   "DB_HMI_ARG1_Seq1_DelaySelect_Blue{4}" : Bool = PLC DB_HMI.ARG1_Seq1_DelaySelect_Blue[4] AT %DB1.DBX0.0, 100 ms
   "DB_HMI_ARG1_Seq1_DelaySelect_Blue{5}" : Bool = PLC DB_HMI.ARG1_Seq1_DelaySelect_Blue[5] AT %DB1.DBX0.0, 100 ms
   "DB_HMI_ARG1_Seq1_DelaySelect_Blue{6}" : Bool = PLC DB_HMI.ARG1_Seq1_DelaySelect_Blue[6] AT %DB1.DBX0.0, 100 ms
   "DB_HMI_ARG1_Seq1_DelaySelect_Blue{7}" : Bool = PLC DB_HMI.ARG1_Seq1_DelaySelect_Blue[7] AT %DB1.DBX0.0, 100 ms
   "DB_HMI_ARG1_Seq1_DelaySelect_Blue{8}" : Bool = PLC DB_HMI.ARG1_Seq1_DelaySelect_Blue[8] AT %DB1.DBX0.0, 100 ms
   "DB_HMI_ARG1_Seq1_DelaySelect_Blue{9}" : Bool = PLC DB_HMI.ARG1_Seq1_DelaySelect_Blue[9] AT %DB1.DBX0.0, 100 ms
   "DB_HMI_ARG1_Seq1_DelaySelect_Blue{10}" : Bool = PLC DB_HMI.ARG1_Seq1_DelaySelect_Blue[10] AT %DB1.DBX0.0, 100 ms
   "DB_HMI_Global_Cmd_Auto" : Bool = PLC DB_HMI.Global_Cmd_Auto, 100 ms
   "DB_HMI_Global_Cmd_Man" : Bool = PLC DB_HMI.Global_Cmd_Man, 100 ms
   "DB_HMI_Global_Cmd_Start" : Bool = PLC DB_HMI.Global_Cmd_Start, 100 ms
   "DB_HMI_Global_Cmd_Stop" : Bool = PLC DB_HMI.Global_Cmd_Stop, 100 ms
   "DB_HMI_Global_Status_Man" : Bool = PLC DB_HMI.Global_Status_Man AT %DB1.DBW0, 100 ms
   "DB_HMI_Global_Status_Auto" : Bool = PLC DB_HMI.Global_Status_Auto AT %DB1.DBW0, 100 ms
   "DB_HMI_Global_selection" : Int = PLC DB_HMI.Global_selection AT %DB1.DBW0, 100 ms
   "DB_HMI_inProduction" : Int = PLC DB_HMI.ARG1_Seq1_inProduction AT %DB1.DBW0, 100 ms

HMI tags "PLC_2_tags"
   "DB_HMI_ARG1_Seq1_S1(1)" : Bool = PLC DB_HMI.ARG1_Seq1_S1, 100 ms
   "DB_HMI_ARG1_Seq1_T1(1)" : Bool = PLC DB_HMI.ARG1_Seq1_T1, 100 ms
   "DB_HMI_ARG1_Seq1_S2(1)" : Bool = PLC DB_HMI.ARG1_Seq1_S2, 100 ms
   "DB_HMI_ARG1_Seq1_T2(1)" : Bool = PLC DB_HMI.ARG1_Seq1_T2, 100 ms
   "DB_HMI_ARG1_Seq1_S3(1)" : Bool = PLC DB_HMI.ARG1_Seq1_S3, 100 ms
   "DB_HMI_ARG1_Seq1_T3(1)" : Bool = PLC DB_HMI.ARG1_Seq1_T3, 100 ms
   "DB_HMI_ARG1_Seq1_S4(1)" : Bool = PLC DB_HMI.ARG1_Seq1_S4, 100 ms
   "DB_HMI_ARG1_Seq1_T4(1)" : Bool = PLC DB_HMI.ARG1_Seq1_T4, 100 ms
   "DB_HMI_ARG1_Seq1_S5(1)" : Bool = PLC DB_HMI.ARG1_Seq1_S5, 100 ms
   "DB_HMI_ARG1_Seq1_T5(1)" : Bool = PLC DB_HMI.ARG1_Seq1_T5, 100 ms
   "DB_HMI_ARG1_Seq1_S6(1)" : Bool = PLC DB_HMI.ARG1_Seq1_S6, 100 ms
   "DB_HMI_ARG1_Seq1_T6(1)" : Bool = PLC DB_HMI.ARG1_Seq1_T6, 100 ms
   "DB_HMI_ARG1_Seq1_S7(1)" : Bool = PLC DB_HMI.ARG1_Seq1_S7, 100 ms
   "DB_HMI_ARG1_Seq1_T7(1)" : Bool = PLC DB_HMI.ARG1_Seq1_T7, 100 ms
   "DB_HMI_ARG1_Seq1_S8(1)" : Bool = PLC DB_HMI.ARG1_Seq1_S8, 100 ms
   "DB_HMI_ARG1_Seq1_T8(1)" : Bool = PLC DB_HMI.ARG1_Seq1_T8, 100 ms
   "DB_HMI_ARG1_Seq1_S9(1)" : Bool = PLC DB_HMI.ARG1_Seq1_S9, 100 ms
   "DB_HMI_ARG1_Seq1_T9(1)" : Bool = PLC DB_HMI.ARG1_Seq1_T9, 100 ms
   "DB_HMI_ARG1_Seq1_S10(1)" : Bool = PLC DB_HMI.ARG1_Seq1_S10, 100 ms
   "DB_HMI_ARG1_Seq1_T10(1)" : Bool = PLC DB_HMI.ARG1_Seq1_T10, 100 ms
   "DB_HMI_ARG1_Seq1_S11(1)" : Bool = PLC DB_HMI.ARG1_Seq1_S11, 100 ms
   "DB_HMI_ARG1_Seq1_T11(1)" : Bool = PLC DB_HMI.ARG1_Seq1_T11, 100 ms
   "DB_HMI_ARG1_Seq1_S12(1)" : Bool = PLC DB_HMI.ARG1_Seq1_S12, 100 ms
   "DB_HMI_ARG1_Seq1_T12(1)" : Bool = PLC DB_HMI.ARG1_Seq1_T12, 100 ms
   "DB_HMI_ARG1_Seq1_S13(1)" : Bool = PLC DB_HMI.ARG1_Seq1_S13, 100 ms
   "DB_HMI_ARG1_Seq1_T13(1)" : Bool = PLC DB_HMI.ARG1_Seq1_T13, 100 ms
   "DB_HMI_ARG1_Seq1_S14(1)" : Bool = PLC DB_HMI.ARG1_Seq1_S14, 100 ms
   "DB_HMI_ARG1_Seq1_T14(1)" : Bool = PLC DB_HMI.ARG1_Seq1_T14, 100 ms
   "DB_HMI_ARG1_Seq1_S15(1)" : Bool = PLC DB_HMI.ARG1_Seq1_S15, 100 ms
   "DB_HMI_ARG1_Seq1_T15(1)" : Bool = PLC DB_HMI.ARG1_Seq1_T15, 100 ms
   "DB_HMI_ARG1_Seq1_S16(1)" : Bool = PLC DB_HMI.ARG1_Seq1_S16, 100 ms
   "DB_HMI_ARG1_Seq1_T16(1)" : Bool = PLC DB_HMI.ARG1_Seq1_T16, 100 ms
   "DB_HMI_ARG1_Seq1_S17(1)" : Bool = PLC DB_HMI.ARG1_Seq1_S17, 100 ms
   "DB_HMI_ARG1_Seq1_T17(1)" : Bool = PLC DB_HMI.ARG1_Seq1_T17, 100 ms
   "DB_HMI_ARG1_Seq1_S18(1)" : Bool = PLC DB_HMI.ARG1_Seq1_S18, 100 ms
   "DB_HMI_ARG1_Seq1_T18(1)" : Bool = PLC DB_HMI.ARG1_Seq1_T18, 100 ms
   "DB_HMI_ARG1_Seq1_S19(1)" : Bool = PLC DB_HMI.ARG1_Seq1_S19, 100 ms
   "DB_HMI_ARG1_Seq1_T19(1)" : Bool = PLC DB_HMI.ARG1_Seq1_T19, 100 ms
   "DB_HMI_inputTimes(1)" : Array [0..8] of DInt = PLC DB_HMI.inputTimes, 100 ms
   "DB_HMI_dropdown_selection(1)" : Int = PLC DB_HMI.dropdown_selection, 100 ms
   "DB_HMI_ARG1_Seq1_Status_Idle(1)" : Bool = PLC DB_HMI.ARG1_Seq1_Status_Idle, 100 ms
   "DB_HMI_ARG1_Seq1_Status_Busy(1)" : Bool = PLC DB_HMI.ARG1_Seq1_Status_Busy, 100 ms
   "DB_HMI_ARG1_Seq1_Status_Man(1)" : Bool = PLC DB_HMI.ARG1_Seq1_Status_Man, 100 ms
   "DB_HMI_ARG1_Seq1_Status_Auto(1)" : Bool = PLC DB_HMI.ARG1_Seq1_Status_Auto, 100 ms
   "DB_HMI_ARG1_Seq1_Cmd_Man(1)" : Bool = PLC DB_HMI.ARG1_Seq1_Cmd_Man, 100 ms
   "DB_HMI_ARG1_Seq1_Cmd_Auto(1)" : Bool = PLC DB_HMI.ARG1_Seq1_Cmd_Auto, 100 ms
   "DB_HMI_ARG1_Seq1_Cmd_Stop(1)" : Bool = PLC DB_HMI.ARG1_Seq1_Cmd_Stop, 100 ms
   "DB_HMI_ARG1_Seq1_Cmd_Start(1)" : Bool = PLC DB_HMI.ARG1_Seq1_Cmd_Start, 100 ms
   "DB_HMI_ARG1_Seq1_Cmd_DelayReset(1)" : Bool = PLC DB_HMI.ARG1_Seq1_Cmd_DelayReset, 100 ms
   "DB_HMI_ARG1_Seq1_Calculated_PT_Red(1)" : Time = PLC DB_HMI.ARG1_Seq1_Calculated_PT_Red, 100 ms
   "DB_HMI_ARG1_Seq1_Calculated_PT_Green(1)" : Time = PLC DB_HMI.ARG1_Seq1_Calculated_PT_Green, 100 ms
   "DB_HMI_ARG1_Seq1_Calculated_PT_Blue(1)" : Time = PLC DB_HMI.ARG1_Seq1_Calculated_PT_Blue, 100 ms
   "DB_HMI_ARG1_Seq1_Messured_PT_Red(1)" : Time = PLC DB_HMI.ARG1_Seq1_Messured_PT_Red, 100 ms
   "DB_HMI_ARG1_Seq1_Messured_PT_Green(1)" : Time = PLC DB_HMI.ARG1_Seq1_Messured_PT_Green, 100 ms
   "DB_HMI_ARG1_Seq1_Messured_PT_Blue(1)" : Time = PLC DB_HMI.ARG1_Seq1_Messured_PT_Blue, 100 ms
   "DB_HMI_ARG1_Seq1_DelaySelect_Red(1)" : Array [0..8] of Bool = PLC DB_HMI.ARG1_Seq1_DelaySelect_Red, 100 ms
   "DB_HMI_ARG1_Seq1_DelaySelect_Green(1)" : Array [0..8] of Bool = PLC DB_HMI.ARG1_Seq1_DelaySelect_Green, 100 ms
   "DB_HMI_ARG1_Seq1_DelaySelect_Blue(1)" : Array [0..8] of Bool = PLC DB_HMI.ARG1_Seq1_DelaySelect_Blue, 100 ms
   "DB_HMI_ARG1_Seq1_DelaySelect_Red{2}(1)" : Bool = PLC DB_HMI.ARG1_Seq1_DelaySelect_Red[2] AT %DB1.DBW0, 100 ms
   "DB_HMI_ARG1_Seq1_DelaySelect_Red{3}(1)" : Bool = PLC DB_HMI.ARG1_Seq1_DelaySelect_Red[3] AT %DB1.DBW0, 100 ms
   "DB_HMI_ARG1_Seq1_DelaySelect_Red{4}(1)" : Bool = PLC DB_HMI.ARG1_Seq1_DelaySelect_Red[4] AT %DB1.DBW0, 100 ms
   "DB_HMI_ARG1_Seq1_DelaySelect_Red{5}(1)" : Bool = PLC DB_HMI.ARG1_Seq1_DelaySelect_Red[5] AT %DB1.DBW0, 100 ms
   "DB_HMI_ARG1_Seq1_DelaySelect_Red{6}(1)" : Bool = PLC DB_HMI.ARG1_Seq1_DelaySelect_Red[6] AT %DB1.DBW0, 100 ms
   "DB_HMI_ARG1_Seq1_DelaySelect_Red{7}(1)" : Bool = PLC DB_HMI.ARG1_Seq1_DelaySelect_Red[7] AT %DB1.DBW0, 100 ms
   "DB_HMI_ARG1_Seq1_DelaySelect_Red{8}(1)" : Bool = PLC DB_HMI.ARG1_Seq1_DelaySelect_Red[8] AT %DB1.DBW0, 100 ms
   "DB_HMI_ARG1_Seq1_DelaySelect_Red{9}(1)" : Bool = PLC DB_HMI.ARG1_Seq1_DelaySelect_Red[9] AT %DB1.DBW0, 100 ms
   "DB_HMI_ARG1_Seq1_DelaySelect_Red{10}(1)" : Bool = PLC DB_HMI.ARG1_Seq1_DelaySelect_Red[10] AT %DB1.DBW0, 100 ms
   "DB_HMI_ARG1_Seq1_DelaySelect_Green{2}(1)" : Bool = PLC DB_HMI.ARG1_Seq1_DelaySelect_Green[2] AT %DB1.DBX0.0, 100 ms
   "DB_HMI_ARG1_Seq1_DelaySelect_Green{3}(1)" : Bool = PLC DB_HMI.ARG1_Seq1_DelaySelect_Green[3] AT %DB1.DBX0.0, 100 ms
   "DB_HMI_ARG1_Seq1_DelaySelect_Green{4}(1)" : Bool = PLC DB_HMI.ARG1_Seq1_DelaySelect_Green[4] AT %DB1.DBX0.0, 100 ms
   "DB_HMI_ARG1_Seq1_DelaySelect_Green{5}(1)" : Bool = PLC DB_HMI.ARG1_Seq1_DelaySelect_Green[5] AT %DB1.DBX0.0, 100 ms
   "DB_HMI_ARG1_Seq1_DelaySelect_Green{6}(1)" : Bool = PLC DB_HMI.ARG1_Seq1_DelaySelect_Green[6] AT %DB1.DBX0.0, 100 ms
   "DB_HMI_ARG1_Seq1_DelaySelect_Green{7}(1)" : Bool = PLC DB_HMI.ARG1_Seq1_DelaySelect_Green[7] AT %DB1.DBX0.0, 100 ms
   "DB_HMI_ARG1_Seq1_DelaySelect_Green{8}(1)" : Bool = PLC DB_HMI.ARG1_Seq1_DelaySelect_Green[8] AT %DB1.DBX0.0, 100 ms
   "DB_HMI_ARG1_Seq1_DelaySelect_Green{9}(1)" : Bool = PLC DB_HMI.ARG1_Seq1_DelaySelect_Green[9] AT %DB1.DBX0.0, 100 ms
   "DB_HMI_ARG1_Seq1_DelaySelect_Green{10}(1)" : Bool = PLC DB_HMI.ARG1_Seq1_DelaySelect_Green[10] AT %DB1.DBX0.0, 100 ms
   "DB_HMI_ARG1_Seq1_DelaySelect_Blue{2}(1)" : Bool = PLC DB_HMI.ARG1_Seq1_DelaySelect_Blue[2] AT %DB1.DBX0.0, 100 ms
   "DB_HMI_ARG1_Seq1_DelaySelect_Blue{3}(1)" : Bool = PLC DB_HMI.ARG1_Seq1_DelaySelect_Blue[3] AT %DB1.DBX0.0, 100 ms
   "DB_HMI_ARG1_Seq1_DelaySelect_Blue{4}(1)" : Bool = PLC DB_HMI.ARG1_Seq1_DelaySelect_Blue[4] AT %DB1.DBX0.0, 100 ms
   "DB_HMI_ARG1_Seq1_DelaySelect_Blue{5}(1)" : Bool = PLC DB_HMI.ARG1_Seq1_DelaySelect_Blue[5] AT %DB1.DBX0.0, 100 ms
   "DB_HMI_ARG1_Seq1_DelaySelect_Blue{6}(1)" : Bool = PLC DB_HMI.ARG1_Seq1_DelaySelect_Blue[6] AT %DB1.DBX0.0, 100 ms
   "DB_HMI_ARG1_Seq1_DelaySelect_Blue{7}(1)" : Bool = PLC DB_HMI.ARG1_Seq1_DelaySelect_Blue[7] AT %DB1.DBX0.0, 100 ms
   "DB_HMI_ARG1_Seq1_DelaySelect_Blue{8}(1)" : Bool = PLC DB_HMI.ARG1_Seq1_DelaySelect_Blue[8] AT %DB1.DBX0.0, 100 ms
   "DB_HMI_ARG1_Seq1_DelaySelect_Blue{9}(1)" : Bool = PLC DB_HMI.ARG1_Seq1_DelaySelect_Blue[9] AT %DB1.DBX0.0, 100 ms
   "DB_HMI_ARG1_Seq1_DelaySelect_Blue{10}(1)" : Bool = PLC DB_HMI.ARG1_Seq1_DelaySelect_Blue[10] AT %DB1.DBX0.0, 100 ms
   "DB_HMI_Global_Cmd_Auto(1)" : Bool = PLC DB_HMI.Global_Cmd_Auto, 100 ms
   "DB_HMI_Global_Cmd_Man(1)" : Bool = PLC DB_HMI.Global_Cmd_Man, 100 ms
   "DB_HMI_Global_Cmd_Start(1)" : Bool = PLC DB_HMI.Global_Cmd_Start, 100 ms
   "DB_HMI_Global_Cmd_Stop(1)" : Bool = PLC DB_HMI.Global_Cmd_Stop, 100 ms
   "DB_HMI_inProduction(1)" : Int = PLC DB_HMI.ARG1_Seq1_inProduction AT %DB1.DBW0, 100 ms

HMI tags "PLC_3_tags"
   "DB_HMI_ARG1_Seq1_S1(2)" : Bool = PLC DB_HMI.ARG1_Seq1_S1, 100 ms
   "DB_HMI_ARG1_Seq1_T1(2)" : Bool = PLC DB_HMI.ARG1_Seq1_T1, 100 ms
   "DB_HMI_ARG1_Seq1_S2(2)" : Bool = PLC DB_HMI.ARG1_Seq1_S2, 100 ms
   "DB_HMI_ARG1_Seq1_T2(2)" : Bool = PLC DB_HMI.ARG1_Seq1_T2, 100 ms
   "DB_HMI_ARG1_Seq1_S3(2)" : Bool = PLC DB_HMI.ARG1_Seq1_S3, 100 ms
   "DB_HMI_ARG1_Seq1_T3(2)" : Bool = PLC DB_HMI.ARG1_Seq1_T3, 100 ms
   "DB_HMI_ARG1_Seq1_S4(2)" : Bool = PLC DB_HMI.ARG1_Seq1_S4, 100 ms
   "DB_HMI_ARG1_Seq1_T4(2)" : Bool = PLC DB_HMI.ARG1_Seq1_T4, 100 ms
   "DB_HMI_ARG1_Seq1_S5(2)" : Bool = PLC DB_HMI.ARG1_Seq1_S5, 100 ms
   "DB_HMI_ARG1_Seq1_T5(2)" : Bool = PLC DB_HMI.ARG1_Seq1_T5, 100 ms
   "DB_HMI_ARG1_Seq1_S6(2)" : Bool = PLC DB_HMI.ARG1_Seq1_S6, 100 ms
   "DB_HMI_ARG1_Seq1_T6(2)" : Bool = PLC DB_HMI.ARG1_Seq1_T6, 100 ms
   "DB_HMI_ARG1_Seq1_S7(2)" : Bool = PLC DB_HMI.ARG1_Seq1_S7, 100 ms
   "DB_HMI_ARG1_Seq1_T7(2)" : Bool = PLC DB_HMI.ARG1_Seq1_T7, 100 ms
   "DB_HMI_ARG1_Seq1_S8(2)" : Bool = PLC DB_HMI.ARG1_Seq1_S8, 100 ms
   "DB_HMI_ARG1_Seq1_T8(2)" : Bool = PLC DB_HMI.ARG1_Seq1_T8, 100 ms
   "DB_HMI_ARG1_Seq1_S9(2)" : Bool = PLC DB_HMI.ARG1_Seq1_S9, 100 ms
   "DB_HMI_ARG1_Seq1_T9(2)" : Bool = PLC DB_HMI.ARG1_Seq1_T9, 100 ms
   "DB_HMI_ARG1_Seq1_S10(2)" : Bool = PLC DB_HMI.ARG1_Seq1_S10, 100 ms
   "DB_HMI_ARG1_Seq1_T10(2)" : Bool = PLC DB_HMI.ARG1_Seq1_T10, 100 ms
   "DB_HMI_ARG1_Seq1_S11(2)" : Bool = PLC DB_HMI.ARG1_Seq1_S11, 100 ms
   "DB_HMI_ARG1_Seq1_T11(2)" : Bool = PLC DB_HMI.ARG1_Seq1_T11, 100 ms
   "DB_HMI_ARG1_Seq1_S12(2)" : Bool = PLC DB_HMI.ARG1_Seq1_S12, 100 ms
   "DB_HMI_ARG1_Seq1_T12(2)" : Bool = PLC DB_HMI.ARG1_Seq1_T12, 100 ms
   "DB_HMI_ARG1_Seq1_S13(2)" : Bool = PLC DB_HMI.ARG1_Seq1_S13, 100 ms
   "DB_HMI_ARG1_Seq1_T13(2)" : Bool = PLC DB_HMI.ARG1_Seq1_T13, 100 ms
   "DB_HMI_ARG1_Seq1_S14(2)" : Bool = PLC DB_HMI.ARG1_Seq1_S14, 100 ms
   "DB_HMI_ARG1_Seq1_T14(2)" : Bool = PLC DB_HMI.ARG1_Seq1_T14, 100 ms
   "DB_HMI_ARG1_Seq1_S15(2)" : Bool = PLC DB_HMI.ARG1_Seq1_S15, 100 ms
   "DB_HMI_ARG1_Seq1_T15(2)" : Bool = PLC DB_HMI.ARG1_Seq1_T15, 100 ms
   "DB_HMI_ARG1_Seq1_S16(2)" : Bool = PLC DB_HMI.ARG1_Seq1_S16, 100 ms
   "DB_HMI_ARG1_Seq1_T16(2)" : Bool = PLC DB_HMI.ARG1_Seq1_T16, 100 ms
   "DB_HMI_ARG1_Seq1_S17(2)" : Bool = PLC DB_HMI.ARG1_Seq1_S17, 100 ms
   "DB_HMI_ARG1_Seq1_T17(2)" : Bool = PLC DB_HMI.ARG1_Seq1_T17, 100 ms
   "DB_HMI_ARG1_Seq1_S18(2)" : Bool = PLC DB_HMI.ARG1_Seq1_S18, 100 ms
   "DB_HMI_ARG1_Seq1_T18(2)" : Bool = PLC DB_HMI.ARG1_Seq1_T18, 100 ms
   "DB_HMI_ARG1_Seq1_S19(2)" : Bool = PLC DB_HMI.ARG1_Seq1_S19, 100 ms
   "DB_HMI_ARG1_Seq1_T19(2)" : Bool = PLC DB_HMI.ARG1_Seq1_T19, 100 ms
   "DB_HMI_inputTimes(2)" : Array [0..8] of DInt = PLC DB_HMI.inputTimes, 100 ms
   "DB_HMI_dropdown_selection(2)" : Int = PLC DB_HMI.dropdown_selection, 100 ms
   "DB_HMI_ARG1_Seq1_Status_Idle(2)" : Bool = PLC DB_HMI.ARG1_Seq1_Status_Idle, 100 ms
   "DB_HMI_ARG1_Seq1_Status_Busy(2)" : Bool = PLC DB_HMI.ARG1_Seq1_Status_Busy, 100 ms
   "DB_HMI_ARG1_Seq1_Status_Man(2)" : Bool = PLC DB_HMI.ARG1_Seq1_Status_Man, 100 ms
   "DB_HMI_ARG1_Seq1_Status_Auto(2)" : Bool = PLC DB_HMI.ARG1_Seq1_Status_Auto, 100 ms
   "DB_HMI_ARG1_Seq1_Cmd_Man(2)" : Bool = PLC DB_HMI.ARG1_Seq1_Cmd_Man, 100 ms
   "DB_HMI_ARG1_Seq1_Cmd_Auto(2)" : Bool = PLC DB_HMI.ARG1_Seq1_Cmd_Auto, 100 ms
   "DB_HMI_ARG1_Seq1_Cmd_Stop(2)" : Bool = PLC DB_HMI.ARG1_Seq1_Cmd_Stop, 100 ms
   "DB_HMI_ARG1_Seq1_Cmd_Start(2)" : Bool = PLC DB_HMI.ARG1_Seq1_Cmd_Start, 100 ms
   "DB_HMI_ARG1_Seq1_Cmd_DelayReset(2)" : Bool = PLC DB_HMI.ARG1_Seq1_Cmd_DelayReset, 100 ms
   "DB_HMI_ARG1_Seq1_Calculated_PT_Red(2)" : Time = PLC DB_HMI.ARG1_Seq1_Calculated_PT_Red, 100 ms
   "DB_HMI_ARG1_Seq1_Calculated_PT_Green(2)" : Time = PLC DB_HMI.ARG1_Seq1_Calculated_PT_Green, 100 ms
   "DB_HMI_ARG1_Seq1_Calculated_PT_Blue(2)" : Time = PLC DB_HMI.ARG1_Seq1_Calculated_PT_Blue, 100 ms
   "DB_HMI_ARG1_Seq1_Messured_PT_Red(2)" : Time = PLC DB_HMI.ARG1_Seq1_Messured_PT_Red, 100 ms
   "DB_HMI_ARG1_Seq1_Messured_PT_Green(2)" : Time = PLC DB_HMI.ARG1_Seq1_Messured_PT_Green, 100 ms
   "DB_HMI_ARG1_Seq1_Messured_PT_Blue(2)" : Time = PLC DB_HMI.ARG1_Seq1_Messured_PT_Blue, 100 ms
   "DB_HMI_ARG1_Seq1_DelaySelect_Red(2)" : Array [0..8] of Bool = PLC DB_HMI.ARG1_Seq1_DelaySelect_Red, 100 ms
   "DB_HMI_ARG1_Seq1_DelaySelect_Green(2)" : Array [0..8] of Bool = PLC DB_HMI.ARG1_Seq1_DelaySelect_Green, 100 ms
   "DB_HMI_ARG1_Seq1_DelaySelect_Blue(2)" : Array [0..8] of Bool = PLC DB_HMI.ARG1_Seq1_DelaySelect_Blue, 100 ms
   "DB_HMI_ARG1_Seq1_DelaySelect_Red{2}(2)" : Bool = PLC DB_HMI.ARG1_Seq1_DelaySelect_Red[2], 100 ms
   "DB_HMI_ARG1_Seq1_DelaySelect_Red{3}(2)" : Bool = PLC DB_HMI.ARG1_Seq1_DelaySelect_Red[3], 100 ms
   "DB_HMI_ARG1_Seq1_DelaySelect_Red{4}(2)" : Bool = PLC DB_HMI.ARG1_Seq1_DelaySelect_Red[4], 100 ms
   "DB_HMI_ARG1_Seq1_DelaySelect_Red{5}(2)" : Bool = PLC DB_HMI.ARG1_Seq1_DelaySelect_Red[5], 100 ms
   "DB_HMI_ARG1_Seq1_DelaySelect_Red{6}(2)" : Bool = PLC DB_HMI.ARG1_Seq1_DelaySelect_Red[6], 100 ms
   "DB_HMI_ARG1_Seq1_DelaySelect_Red{7}(2)" : Bool = PLC DB_HMI.ARG1_Seq1_DelaySelect_Red[7], 100 ms
   "DB_HMI_ARG1_Seq1_DelaySelect_Red{8}(2)" : Bool = PLC DB_HMI.ARG1_Seq1_DelaySelect_Red[8], 100 ms
   "DB_HMI_ARG1_Seq1_DelaySelect_Red{9}(2)" : Bool = PLC DB_HMI.ARG1_Seq1_DelaySelect_Red[9], 100 ms
   "DB_HMI_ARG1_Seq1_DelaySelect_Red{10}(2)" : Bool = PLC DB_HMI.ARG1_Seq1_DelaySelect_Red[10], 100 ms
   "DB_HMI_ARG1_Seq1_DelaySelect_Green{2}(2)" : Bool = PLC DB_HMI.ARG1_Seq1_DelaySelect_Green[2], 100 ms
   "DB_HMI_ARG1_Seq1_DelaySelect_Green{3}(2)" : Bool = PLC DB_HMI.ARG1_Seq1_DelaySelect_Green[3], 100 ms
   "DB_HMI_ARG1_Seq1_DelaySelect_Green{4}(2)" : Bool = PLC DB_HMI.ARG1_Seq1_DelaySelect_Green[4], 100 ms
   "DB_HMI_ARG1_Seq1_DelaySelect_Green{5}(2)" : Bool = PLC DB_HMI.ARG1_Seq1_DelaySelect_Green[5], 100 ms
   "DB_HMI_ARG1_Seq1_DelaySelect_Green{6}(2)" : Bool = PLC DB_HMI.ARG1_Seq1_DelaySelect_Green[6], 100 ms
   "DB_HMI_ARG1_Seq1_DelaySelect_Green{7}(2)" : Bool = PLC DB_HMI.ARG1_Seq1_DelaySelect_Green[7], 100 ms
   "DB_HMI_ARG1_Seq1_DelaySelect_Green{8}(2)" : Bool = PLC DB_HMI.ARG1_Seq1_DelaySelect_Green[8], 100 ms
   "DB_HMI_ARG1_Seq1_DelaySelect_Green{9}(2)" : Bool = PLC DB_HMI.ARG1_Seq1_DelaySelect_Green[9], 100 ms
   "DB_HMI_ARG1_Seq1_DelaySelect_Green{10}(2)" : Bool = PLC DB_HMI.ARG1_Seq1_DelaySelect_Green[10], 100 ms
   "DB_HMI_ARG1_Seq1_DelaySelect_Blue{2}(2)" : Bool = PLC DB_HMI.ARG1_Seq1_DelaySelect_Blue[2], 100 ms
   "DB_HMI_ARG1_Seq1_DelaySelect_Blue{3}(2)" : Bool = PLC DB_HMI.ARG1_Seq1_DelaySelect_Blue[3], 100 ms
   "DB_HMI_ARG1_Seq1_DelaySelect_Blue{4}(2)" : Bool = PLC DB_HMI.ARG1_Seq1_DelaySelect_Blue[4], 100 ms
   "DB_HMI_ARG1_Seq1_DelaySelect_Blue{5}(2)" : Bool = PLC DB_HMI.ARG1_Seq1_DelaySelect_Blue[5], 100 ms
   "DB_HMI_ARG1_Seq1_DelaySelect_Blue{6}(2)" : Bool = PLC DB_HMI.ARG1_Seq1_DelaySelect_Blue[6], 100 ms
   "DB_HMI_ARG1_Seq1_DelaySelect_Blue{7}(2)" : Bool = PLC DB_HMI.ARG1_Seq1_DelaySelect_Blue[7], 100 ms
   "DB_HMI_ARG1_Seq1_DelaySelect_Blue{8}(2)" : Bool = PLC DB_HMI.ARG1_Seq1_DelaySelect_Blue[8], 100 ms
   "DB_HMI_ARG1_Seq1_DelaySelect_Blue{9}(2)" : Bool = PLC DB_HMI.ARG1_Seq1_DelaySelect_Blue[9], 100 ms
   "DB_HMI_ARG1_Seq1_DelaySelect_Blue{10}(2)" : Bool = PLC DB_HMI.ARG1_Seq1_DelaySelect_Blue[10], 100 ms
   "DB_HMI_Global_Cmd_Auto(2)" : Bool = PLC DB_HMI.Global_Cmd_Auto, 100 ms
   "DB_HMI_Global_Cmd_Man(2)" : Bool = PLC DB_HMI.Global_Cmd_Man, 100 ms
   "DB_HMI_Global_Cmd_Start(2)" : Bool = PLC DB_HMI.Global_Cmd_Start, 100 ms
   "DB_HMI_Global_Cmd_Stop(2)" : Bool = PLC DB_HMI.Global_Cmd_Stop, 100 ms
   "DB_HMI_inProduction(2)" : Int = PLC DB_HMI.ARG1_Seq1_inProduction AT %DB1.DBW0, 100 ms

HMI tags "PLC_4_tags"
   "DB_HMI_ARG1_Seq1_S1(3)" : Bool = PLC DB_HMI.ARG1_Seq1_S1, 100 ms
   "DB_HMI_ARG1_Seq1_T1(3)" : Bool = PLC DB_HMI.ARG1_Seq1_T1, 100 ms
   "DB_HMI_ARG1_Seq1_S2(3)" : Bool = PLC DB_HMI.ARG1_Seq1_S2, 100 ms
   "DB_HMI_ARG1_Seq1_T2(3)" : Bool = PLC DB_HMI.ARG1_Seq1_T2, 100 ms
   "DB_HMI_ARG1_Seq1_S3(3)" : Bool = PLC DB_HMI.ARG1_Seq1_S3, 100 ms
   "DB_HMI_ARG1_Seq1_T3(3)" : Bool = PLC DB_HMI.ARG1_Seq1_T3, 100 ms
   "DB_HMI_ARG1_Seq1_S4(3)" : Bool = PLC DB_HMI.ARG1_Seq1_S4, 100 ms
   "DB_HMI_ARG1_Seq1_T4(3)" : Bool = PLC DB_HMI.ARG1_Seq1_T4, 100 ms
   "DB_HMI_ARG1_Seq1_S5(3)" : Bool = PLC DB_HMI.ARG1_Seq1_S5, 100 ms
   "DB_HMI_ARG1_Seq1_T5(3)" : Bool = PLC DB_HMI.ARG1_Seq1_T5, 100 ms
   "DB_HMI_ARG1_Seq1_S6(3)" : Bool = PLC DB_HMI.ARG1_Seq1_S6, 100 ms
   "DB_HMI_ARG1_Seq1_T6(3)" : Bool = PLC DB_HMI.ARG1_Seq1_T6, 100 ms
   "DB_HMI_ARG1_Seq1_S7(3)" : Bool = PLC DB_HMI.ARG1_Seq1_S7, 100 ms
   "DB_HMI_ARG1_Seq1_T7(3)" : Bool = PLC DB_HMI.ARG1_Seq1_T7, 100 ms
   "DB_HMI_ARG1_Seq1_S8(3)" : Bool = PLC DB_HMI.ARG1_Seq1_S8, 100 ms
   "DB_HMI_ARG1_Seq1_T8(3)" : Bool = PLC DB_HMI.ARG1_Seq1_T8, 100 ms
   "DB_HMI_ARG1_Seq1_S9(3)" : Bool = PLC DB_HMI.ARG1_Seq1_S9, 100 ms
   "DB_HMI_ARG1_Seq1_T9(3)" : Bool = PLC DB_HMI.ARG1_Seq1_T9, 100 ms
   "DB_HMI_ARG1_Seq1_S10(3)" : Bool = PLC DB_HMI.ARG1_Seq1_S10, 100 ms
   "DB_HMI_ARG1_Seq1_T10(3)" : Bool = PLC DB_HMI.ARG1_Seq1_T10, 100 ms
   "DB_HMI_ARG1_Seq1_S11(3)" : Bool = PLC DB_HMI.ARG1_Seq1_S11, 100 ms
   "DB_HMI_ARG1_Seq1_T11(3)" : Bool = PLC DB_HMI.ARG1_Seq1_T11, 100 ms
   "DB_HMI_ARG1_Seq1_S12(3)" : Bool = PLC DB_HMI.ARG1_Seq1_S12, 100 ms
   "DB_HMI_ARG1_Seq1_T12(3)" : Bool = PLC DB_HMI.ARG1_Seq1_T12, 100 ms
   "DB_HMI_ARG1_Seq1_S13(3)" : Bool = PLC DB_HMI.ARG1_Seq1_S13, 100 ms
   "DB_HMI_ARG1_Seq1_T13(3)" : Bool = PLC DB_HMI.ARG1_Seq1_T13, 100 ms
   "DB_HMI_ARG1_Seq1_S14(3)" : Bool = PLC DB_HMI.ARG1_Seq1_S14, 100 ms
   "DB_HMI_ARG1_Seq1_T14(3)" : Bool = PLC DB_HMI.ARG1_Seq1_T14, 100 ms
   "DB_HMI_ARG1_Seq1_S15(3)" : Bool = PLC DB_HMI.ARG1_Seq1_S15, 100 ms
   "DB_HMI_ARG1_Seq1_T15(3)" : Bool = PLC DB_HMI.ARG1_Seq1_T15, 100 ms
   "DB_HMI_ARG1_Seq1_S16(3)" : Bool = PLC DB_HMI.ARG1_Seq1_S16, 100 ms
   "DB_HMI_ARG1_Seq1_T16(3)" : Bool = PLC DB_HMI.ARG1_Seq1_T16, 100 ms
   "DB_HMI_ARG1_Seq1_S17(3)" : Bool = PLC DB_HMI.ARG1_Seq1_S17, 100 ms
   "DB_HMI_ARG1_Seq1_T17(3)" : Bool = PLC DB_HMI.ARG1_Seq1_T17, 100 ms
   "DB_HMI_ARG1_Seq1_S18(3)" : Bool = PLC DB_HMI.ARG1_Seq1_S18, 100 ms
   "DB_HMI_ARG1_Seq1_T18(3)" : Bool = PLC DB_HMI.ARG1_Seq1_T18, 100 ms
   "DB_HMI_ARG1_Seq1_S19(3)" : Bool = PLC DB_HMI.ARG1_Seq1_S19, 100 ms
   "DB_HMI_ARG1_Seq1_T19(3)" : Bool = PLC DB_HMI.ARG1_Seq1_T19, 100 ms
   "DB_HMI_inputTimes(3)" : Array [0..8] of DInt = PLC DB_HMI.inputTimes, 100 ms
   "DB_HMI_dropdown_selection(3)" : Int = PLC DB_HMI.dropdown_selection, 100 ms
   "DB_HMI_ARG1_Seq1_Status_Idle(3)" : Bool = PLC DB_HMI.ARG1_Seq1_Status_Idle, 100 ms
   "DB_HMI_ARG1_Seq1_Status_Busy(3)" : Bool = PLC DB_HMI.ARG1_Seq1_Status_Busy, 100 ms
   "DB_HMI_ARG1_Seq1_Status_Man(3)" : Bool = PLC DB_HMI.ARG1_Seq1_Status_Man, 100 ms
   "DB_HMI_ARG1_Seq1_Status_Auto(3)" : Bool = PLC DB_HMI.ARG1_Seq1_Status_Auto, 100 ms
   "DB_HMI_ARG1_Seq1_Cmd_Man(3)" : Bool = PLC DB_HMI.ARG1_Seq1_Cmd_Man, 100 ms
   "DB_HMI_ARG1_Seq1_Cmd_Auto(3)" : Bool = PLC DB_HMI.ARG1_Seq1_Cmd_Auto, 100 ms
   "DB_HMI_ARG1_Seq1_Cmd_Stop(3)" : Bool = PLC DB_HMI.ARG1_Seq1_Cmd_Stop, 100 ms
   "DB_HMI_ARG1_Seq1_Cmd_Start(3)" : Bool = PLC DB_HMI.ARG1_Seq1_Cmd_Start, 100 ms
   "DB_HMI_ARG1_Seq1_Cmd_DelayReset(3)" : Bool = PLC DB_HMI.ARG1_Seq1_Cmd_DelayReset, 100 ms
   "DB_HMI_ARG1_Seq1_Calculated_PT_Red(3)" : Time = PLC DB_HMI.ARG1_Seq1_Calculated_PT_Red, 100 ms
   "DB_HMI_ARG1_Seq1_Calculated_PT_Green(3)" : Time = PLC DB_HMI.ARG1_Seq1_Calculated_PT_Green, 100 ms
   "DB_HMI_ARG1_Seq1_Calculated_PT_Blue(3)" : Time = PLC DB_HMI.ARG1_Seq1_Calculated_PT_Blue, 100 ms
   "DB_HMI_ARG1_Seq1_Messured_PT_Red(3)" : Time = PLC DB_HMI.ARG1_Seq1_Messured_PT_Red, 100 ms
   "DB_HMI_ARG1_Seq1_Messured_PT_Green(3)" : Time = PLC DB_HMI.ARG1_Seq1_Messured_PT_Green, 100 ms
   "DB_HMI_ARG1_Seq1_Messured_PT_Blue(3)" : Time = PLC DB_HMI.ARG1_Seq1_Messured_PT_Blue, 100 ms
   "DB_HMI_ARG1_Seq1_DelaySelect_Red(3)" : Array [0..8] of Bool = PLC DB_HMI.ARG1_Seq1_DelaySelect_Red, 100 ms
   "DB_HMI_ARG1_Seq1_DelaySelect_Green(3)" : Array [0..8] of Bool = PLC DB_HMI.ARG1_Seq1_DelaySelect_Green, 100 ms
   "DB_HMI_ARG1_Seq1_DelaySelect_Blue(3)" : Array [0..8] of Bool = PLC DB_HMI.ARG1_Seq1_DelaySelect_Blue, 100 ms
   "DB_HMI_ARG1_Seq1_DelaySelect_Red{2}(3)" : Bool = PLC DB_HMI.ARG1_Seq1_DelaySelect_Red[2], 100 ms
   "DB_HMI_ARG1_Seq1_DelaySelect_Red{3}(3)" : Bool = PLC DB_HMI.ARG1_Seq1_DelaySelect_Red[3], 100 ms
   "DB_HMI_ARG1_Seq1_DelaySelect_Red{4}(3)" : Bool = PLC DB_HMI.ARG1_Seq1_DelaySelect_Red[4], 100 ms
   "DB_HMI_ARG1_Seq1_DelaySelect_Red{5}(3)" : Bool = PLC DB_HMI.ARG1_Seq1_DelaySelect_Red[5], 100 ms
   "DB_HMI_ARG1_Seq1_DelaySelect_Red{6}(3)" : Bool = PLC DB_HMI.ARG1_Seq1_DelaySelect_Red[6], 100 ms
   "DB_HMI_ARG1_Seq1_DelaySelect_Red{7}(3)" : Bool = PLC DB_HMI.ARG1_Seq1_DelaySelect_Red[7], 100 ms
   "DB_HMI_ARG1_Seq1_DelaySelect_Red{8}(3)" : Bool = PLC DB_HMI.ARG1_Seq1_DelaySelect_Red[8], 100 ms
   "DB_HMI_ARG1_Seq1_DelaySelect_Red{9}(3)" : Bool = PLC DB_HMI.ARG1_Seq1_DelaySelect_Red[9], 100 ms
   "DB_HMI_ARG1_Seq1_DelaySelect_Red{10}(3)" : Bool = PLC DB_HMI.ARG1_Seq1_DelaySelect_Red[10], 100 ms
   "DB_HMI_ARG1_Seq1_DelaySelect_Green{2}(3)" : Bool = PLC DB_HMI.ARG1_Seq1_DelaySelect_Green[2], 100 ms
   "DB_HMI_ARG1_Seq1_DelaySelect_Green{3}(3)" : Bool = PLC DB_HMI.ARG1_Seq1_DelaySelect_Green[3], 100 ms
   "DB_HMI_ARG1_Seq1_DelaySelect_Green{4}(3)" : Bool = PLC DB_HMI.ARG1_Seq1_DelaySelect_Green[4], 100 ms
   "DB_HMI_ARG1_Seq1_DelaySelect_Green{5}(3)" : Bool = PLC DB_HMI.ARG1_Seq1_DelaySelect_Green[5], 100 ms
   "DB_HMI_ARG1_Seq1_DelaySelect_Green{6}(3)" : Bool = PLC DB_HMI.ARG1_Seq1_DelaySelect_Green[6], 100 ms
   "DB_HMI_ARG1_Seq1_DelaySelect_Green{7}(3)" : Bool = PLC DB_HMI.ARG1_Seq1_DelaySelect_Green[7], 100 ms
   "DB_HMI_ARG1_Seq1_DelaySelect_Green{8}(3)" : Bool = PLC DB_HMI.ARG1_Seq1_DelaySelect_Green[8], 100 ms
   "DB_HMI_ARG1_Seq1_DelaySelect_Green{9}(3)" : Bool = PLC DB_HMI.ARG1_Seq1_DelaySelect_Green[9], 100 ms
   "DB_HMI_ARG1_Seq1_DelaySelect_Green{10}(3)" : Bool = PLC DB_HMI.ARG1_Seq1_DelaySelect_Green[10], 100 ms
   "DB_HMI_ARG1_Seq1_DelaySelect_Blue{2}(3)" : Bool = PLC DB_HMI.ARG1_Seq1_DelaySelect_Blue[2], 100 ms
   "DB_HMI_ARG1_Seq1_DelaySelect_Blue{3}(3)" : Bool = PLC DB_HMI.ARG1_Seq1_DelaySelect_Blue[3], 100 ms
   "DB_HMI_ARG1_Seq1_DelaySelect_Blue{4}(3)" : Bool = PLC DB_HMI.ARG1_Seq1_DelaySelect_Blue[4], 100 ms
   "DB_HMI_ARG1_Seq1_DelaySelect_Blue{5}(3)" : Bool = PLC DB_HMI.ARG1_Seq1_DelaySelect_Blue[5], 100 ms
   "DB_HMI_ARG1_Seq1_DelaySelect_Blue{6}(3)" : Bool = PLC DB_HMI.ARG1_Seq1_DelaySelect_Blue[6], 100 ms
   "DB_HMI_ARG1_Seq1_DelaySelect_Blue{7}(3)" : Bool = PLC DB_HMI.ARG1_Seq1_DelaySelect_Blue[7], 100 ms
   "DB_HMI_ARG1_Seq1_DelaySelect_Blue{8}(3)" : Bool = PLC DB_HMI.ARG1_Seq1_DelaySelect_Blue[8], 100 ms
   "DB_HMI_ARG1_Seq1_DelaySelect_Blue{9}(3)" : Bool = PLC DB_HMI.ARG1_Seq1_DelaySelect_Blue[9], 100 ms
   "DB_HMI_ARG1_Seq1_DelaySelect_Blue{10}(3)" : Bool = PLC DB_HMI.ARG1_Seq1_DelaySelect_Blue[10], 100 ms
   "DB_HMI_Global_Cmd_Auto(3)" : Bool = PLC DB_HMI.Global_Cmd_Auto, 100 ms
   "DB_HMI_Global_Cmd_Man(3)" : Bool = PLC DB_HMI.Global_Cmd_Man, 100 ms
   "DB_HMI_Global_Cmd_Start(3)" : Bool = PLC DB_HMI.Global_Cmd_Start, 100 ms
   "DB_HMI_Global_Cmd_Stop(3)" : Bool = PLC DB_HMI.Global_Cmd_Stop, 100 ms
   "DB_HMI_inProduction(3)" : Int = PLC DB_HMI.ARG1_Seq1_inProduction AT %DB1.DBW0, 100 ms

HMI tags "PLC_5_tags"
   "DB_HMI_ARG1_Seq1_S1(4)" : Bool = PLC DB_HMI.ARG1_Seq1_S1, 100 ms
   "DB_HMI_ARG1_Seq1_T1(4)" : Bool = PLC DB_HMI.ARG1_Seq1_T1, 100 ms
   "DB_HMI_ARG1_Seq1_S2(4)" : Bool = PLC DB_HMI.ARG1_Seq1_S2, 100 ms
   "DB_HMI_ARG1_Seq1_T2(4)" : Bool = PLC DB_HMI.ARG1_Seq1_T2, 100 ms
   "DB_HMI_ARG1_Seq1_S3(4)" : Bool = PLC DB_HMI.ARG1_Seq1_S3, 100 ms
   "DB_HMI_ARG1_Seq1_T3(4)" : Bool = PLC DB_HMI.ARG1_Seq1_T3, 100 ms
   "DB_HMI_ARG1_Seq1_S4(4)" : Bool = PLC DB_HMI.ARG1_Seq1_S4, 100 ms
   "DB_HMI_ARG1_Seq1_T4(4)" : Bool = PLC DB_HMI.ARG1_Seq1_T4, 100 ms
   "DB_HMI_ARG1_Seq1_S5(4)" : Bool = PLC DB_HMI.ARG1_Seq1_S5, 100 ms
   "DB_HMI_ARG1_Seq1_T5(4)" : Bool = PLC DB_HMI.ARG1_Seq1_T5, 100 ms
   "DB_HMI_ARG1_Seq1_S6(4)" : Bool = PLC DB_HMI.ARG1_Seq1_S6, 100 ms
   "DB_HMI_ARG1_Seq1_T6(4)" : Bool = PLC DB_HMI.ARG1_Seq1_T6, 100 ms
   "DB_HMI_ARG1_Seq1_S7(4)" : Bool = PLC DB_HMI.ARG1_Seq1_S7, 100 ms
   "DB_HMI_ARG1_Seq1_T7(4)" : Bool = PLC DB_HMI.ARG1_Seq1_T7, 100 ms
   "DB_HMI_ARG1_Seq1_S8(4)" : Bool = PLC DB_HMI.ARG1_Seq1_S8, 100 ms
   "DB_HMI_ARG1_Seq1_T8(4)" : Bool = PLC DB_HMI.ARG1_Seq1_T8, 100 ms
   "DB_HMI_ARG1_Seq1_S9(4)" : Bool = PLC DB_HMI.ARG1_Seq1_S9, 100 ms
   "DB_HMI_ARG1_Seq1_T9(4)" : Bool = PLC DB_HMI.ARG1_Seq1_T9, 100 ms
   "DB_HMI_ARG1_Seq1_S10(4)" : Bool = PLC DB_HMI.ARG1_Seq1_S10, 100 ms
   "DB_HMI_ARG1_Seq1_T10(4)" : Bool = PLC DB_HMI.ARG1_Seq1_T10, 100 ms
   "DB_HMI_ARG1_Seq1_S11(4)" : Bool = PLC DB_HMI.ARG1_Seq1_S11, 100 ms
   "DB_HMI_ARG1_Seq1_T11(4)" : Bool = PLC DB_HMI.ARG1_Seq1_T11, 100 ms
   "DB_HMI_ARG1_Seq1_S12(4)" : Bool = PLC DB_HMI.ARG1_Seq1_S12, 100 ms
   "DB_HMI_ARG1_Seq1_T12(4)" : Bool = PLC DB_HMI.ARG1_Seq1_T12, 100 ms
   "DB_HMI_ARG1_Seq1_S13(4)" : Bool = PLC DB_HMI.ARG1_Seq1_S13, 100 ms
   "DB_HMI_ARG1_Seq1_T13(4)" : Bool = PLC DB_HMI.ARG1_Seq1_T13, 100 ms
   "DB_HMI_ARG1_Seq1_S14(4)" : Bool = PLC DB_HMI.ARG1_Seq1_S14, 100 ms
   "DB_HMI_ARG1_Seq1_T14(4)" : Bool = PLC DB_HMI.ARG1_Seq1_T14, 100 ms
   "DB_HMI_ARG1_Seq1_S15(4)" : Bool = PLC DB_HMI.ARG1_Seq1_S15, 100 ms
   "DB_HMI_ARG1_Seq1_T15(4)" : Bool = PLC DB_HMI.ARG1_Seq1_T15, 100 ms
   "DB_HMI_ARG1_Seq1_S16(4)" : Bool = PLC DB_HMI.ARG1_Seq1_S16, 100 ms
   "DB_HMI_ARG1_Seq1_T16(4)" : Bool = PLC DB_HMI.ARG1_Seq1_T16, 100 ms
   "DB_HMI_ARG1_Seq1_S17(4)" : Bool = PLC DB_HMI.ARG1_Seq1_S17, 100 ms
   "DB_HMI_ARG1_Seq1_T17(4)" : Bool = PLC DB_HMI.ARG1_Seq1_T17, 100 ms
   "DB_HMI_ARG1_Seq1_S18(4)" : Bool = PLC DB_HMI.ARG1_Seq1_S18, 100 ms
   "DB_HMI_ARG1_Seq1_T18(4)" : Bool = PLC DB_HMI.ARG1_Seq1_T18, 100 ms
   "DB_HMI_ARG1_Seq1_S19(4)" : Bool = PLC DB_HMI.ARG1_Seq1_S19, 100 ms
   "DB_HMI_ARG1_Seq1_T19(4)" : Bool = PLC DB_HMI.ARG1_Seq1_T19, 100 ms
   "DB_HMI_inputTimes(4)" : Array [0..8] of DInt = PLC DB_HMI.inputTimes, 100 ms
   "DB_HMI_dropdown_selection(4)" : Int = PLC DB_HMI.dropdown_selection, 100 ms
   "DB_HMI_ARG1_Seq1_Status_Idle(4)" : Bool = PLC DB_HMI.ARG1_Seq1_Status_Idle, 100 ms
   "DB_HMI_ARG1_Seq1_Status_Busy(4)" : Bool = PLC DB_HMI.ARG1_Seq1_Status_Busy, 100 ms
   "DB_HMI_ARG1_Seq1_Status_Man(4)" : Bool = PLC DB_HMI.ARG1_Seq1_Status_Man, 100 ms
   "DB_HMI_ARG1_Seq1_Status_Auto(4)" : Bool = PLC DB_HMI.ARG1_Seq1_Status_Auto, 100 ms
   "DB_HMI_ARG1_Seq1_Cmd_Man(4)" : Bool = PLC DB_HMI.ARG1_Seq1_Cmd_Man, 100 ms
   "DB_HMI_ARG1_Seq1_Cmd_Auto(4)" : Bool = PLC DB_HMI.ARG1_Seq1_Cmd_Auto, 100 ms
   "DB_HMI_ARG1_Seq1_Cmd_Stop(4)" : Bool = PLC DB_HMI.ARG1_Seq1_Cmd_Stop, 100 ms
   "DB_HMI_ARG1_Seq1_Cmd_Start(4)" : Bool = PLC DB_HMI.ARG1_Seq1_Cmd_Start, 100 ms
   "DB_HMI_ARG1_Seq1_Cmd_DelayReset(4)" : Bool = PLC DB_HMI.ARG1_Seq1_Cmd_DelayReset, 100 ms
   "DB_HMI_ARG1_Seq1_Calculated_PT_Red(4)" : Time = PLC DB_HMI.ARG1_Seq1_Calculated_PT_Red, 100 ms
   "DB_HMI_ARG1_Seq1_Calculated_PT_Green(4)" : Time = PLC DB_HMI.ARG1_Seq1_Calculated_PT_Green, 100 ms
   "DB_HMI_ARG1_Seq1_Calculated_PT_Blue(4)" : Time = PLC DB_HMI.ARG1_Seq1_Calculated_PT_Blue, 100 ms
   "DB_HMI_ARG1_Seq1_Messured_PT_Red(4)" : Time = PLC DB_HMI.ARG1_Seq1_Messured_PT_Red, 100 ms
   "DB_HMI_ARG1_Seq1_Messured_PT_Green(4)" : Time = PLC DB_HMI.ARG1_Seq1_Messured_PT_Green, 100 ms
   "DB_HMI_ARG1_Seq1_Messured_PT_Blue(4)" : Time = PLC DB_HMI.ARG1_Seq1_Messured_PT_Blue, 100 ms
   "DB_HMI_ARG1_Seq1_DelaySelect_Red(4)" : Array [0..8] of Bool = PLC DB_HMI.ARG1_Seq1_DelaySelect_Red, 100 ms
   "DB_HMI_ARG1_Seq1_DelaySelect_Green(4)" : Array [0..8] of Bool = PLC DB_HMI.ARG1_Seq1_DelaySelect_Green, 100 ms
   "DB_HMI_ARG1_Seq1_DelaySelect_Blue(4)" : Array [0..8] of Bool = PLC DB_HMI.ARG1_Seq1_DelaySelect_Blue, 100 ms
   "DB_HMI_ARG1_Seq1_DelaySelect_Red{2}(4)" : Bool = PLC DB_HMI.ARG1_Seq1_DelaySelect_Red[2], 100 ms
   "DB_HMI_ARG1_Seq1_DelaySelect_Red{3}(4)" : Bool = PLC DB_HMI.ARG1_Seq1_DelaySelect_Red[3], 100 ms
   "DB_HMI_ARG1_Seq1_DelaySelect_Red{4}(4)" : Bool = PLC DB_HMI.ARG1_Seq1_DelaySelect_Red[4], 100 ms
   "DB_HMI_ARG1_Seq1_DelaySelect_Red{5}(4)" : Bool = PLC DB_HMI.ARG1_Seq1_DelaySelect_Red[5], 100 ms
   "DB_HMI_ARG1_Seq1_DelaySelect_Red{6}(4)" : Bool = PLC DB_HMI.ARG1_Seq1_DelaySelect_Red[6], 100 ms
   "DB_HMI_ARG1_Seq1_DelaySelect_Red{7}(4)" : Bool = PLC DB_HMI.ARG1_Seq1_DelaySelect_Red[7], 100 ms
   "DB_HMI_ARG1_Seq1_DelaySelect_Red{8}(4)" : Bool = PLC DB_HMI.ARG1_Seq1_DelaySelect_Red[8], 100 ms
   "DB_HMI_ARG1_Seq1_DelaySelect_Red{9}(4)" : Bool = PLC DB_HMI.ARG1_Seq1_DelaySelect_Red[9], 100 ms
   "DB_HMI_ARG1_Seq1_DelaySelect_Red{10}(4)" : Bool = PLC DB_HMI.ARG1_Seq1_DelaySelect_Red[10], 100 ms
   "DB_HMI_ARG1_Seq1_DelaySelect_Green{2}(4)" : Bool = PLC DB_HMI.ARG1_Seq1_DelaySelect_Green[2], 100 ms
   "DB_HMI_ARG1_Seq1_DelaySelect_Green{3}(4)" : Bool = PLC DB_HMI.ARG1_Seq1_DelaySelect_Green[3], 100 ms
   "DB_HMI_ARG1_Seq1_DelaySelect_Green{4}(4)" : Bool = PLC DB_HMI.ARG1_Seq1_DelaySelect_Green[4], 100 ms
   "DB_HMI_ARG1_Seq1_DelaySelect_Green{5}(4)" : Bool = PLC DB_HMI.ARG1_Seq1_DelaySelect_Green[5], 100 ms
   "DB_HMI_ARG1_Seq1_DelaySelect_Green{6}(4)" : Bool = PLC DB_HMI.ARG1_Seq1_DelaySelect_Green[6], 100 ms
   "DB_HMI_ARG1_Seq1_DelaySelect_Green{7}(4)" : Bool = PLC DB_HMI.ARG1_Seq1_DelaySelect_Green[7], 100 ms
   "DB_HMI_ARG1_Seq1_DelaySelect_Green{8}(4)" : Bool = PLC DB_HMI.ARG1_Seq1_DelaySelect_Green[8], 100 ms
   "DB_HMI_ARG1_Seq1_DelaySelect_Green{9}(4)" : Bool = PLC DB_HMI.ARG1_Seq1_DelaySelect_Green[9], 100 ms
   "DB_HMI_ARG1_Seq1_DelaySelect_Green{10}(4)" : Bool = PLC DB_HMI.ARG1_Seq1_DelaySelect_Green[10], 100 ms
   "DB_HMI_ARG1_Seq1_DelaySelect_Blue{2}(4)" : Bool = PLC DB_HMI.ARG1_Seq1_DelaySelect_Blue[2], 100 ms
   "DB_HMI_ARG1_Seq1_DelaySelect_Blue{3}(4)" : Bool = PLC DB_HMI.ARG1_Seq1_DelaySelect_Blue[3], 100 ms
   "DB_HMI_ARG1_Seq1_DelaySelect_Blue{4}(4)" : Bool = PLC DB_HMI.ARG1_Seq1_DelaySelect_Blue[4], 100 ms
   "DB_HMI_ARG1_Seq1_DelaySelect_Blue{5}(4)" : Bool = PLC DB_HMI.ARG1_Seq1_DelaySelect_Blue[5], 100 ms
   "DB_HMI_ARG1_Seq1_DelaySelect_Blue{6}(4)" : Bool = PLC DB_HMI.ARG1_Seq1_DelaySelect_Blue[6], 100 ms
   "DB_HMI_ARG1_Seq1_DelaySelect_Blue{7}(4)" : Bool = PLC DB_HMI.ARG1_Seq1_DelaySelect_Blue[7], 100 ms
   "DB_HMI_ARG1_Seq1_DelaySelect_Blue{8}(4)" : Bool = PLC DB_HMI.ARG1_Seq1_DelaySelect_Blue[8], 100 ms
   "DB_HMI_ARG1_Seq1_DelaySelect_Blue{9}(4)" : Bool = PLC DB_HMI.ARG1_Seq1_DelaySelect_Blue[9], 100 ms
   "DB_HMI_ARG1_Seq1_DelaySelect_Blue{10}(4)" : Bool = PLC DB_HMI.ARG1_Seq1_DelaySelect_Blue[10], 100 ms
   "DB_HMI_Global_Cmd_Auto(4)" : Bool = PLC DB_HMI.Global_Cmd_Auto, 100 ms
   "DB_HMI_Global_Cmd_Man(4)" : Bool = PLC DB_HMI.Global_Cmd_Man, 100 ms
   "DB_HMI_Global_Cmd_Start(4)" : Bool = PLC DB_HMI.Global_Cmd_Start, 100 ms
   "DB_HMI_Global_Cmd_Stop(4)" : Bool = PLC DB_HMI.Global_Cmd_Stop, 100 ms
   "DB_HMI_inProduction(4)" : Int = PLC DB_HMI.ARG1_Seq1_inProduction AT %DB1.DBW0, 100 ms

HMI tags "Template"
   "MainNavigationState" : Int, internal
   "SubNavigationState" : Int, internal
   "CurrentUserName" : WString[18], internal
   "DiagState" : Int, internal
   "PopUpBackground" : Bool, internal
   "UserName" : WString[20], internal
   "Password" : WString[20], internal
   "UserIsLoggedIn" : Bool, internal
   "CodeView" : Bool, internal
   "Brightness" : Int, internal
      on ChangeValue: function_e4c2bb66("Brightness")
   "CurrentLanguage" : Bool, internal
   "CurrentRecipeName" : WString[30], internal
   "CurrentMachineState" : Int, internal
   "OptionPanelNavigationState" : Int, internal
   "ButtonDown" : Bool, internal
   "ThirdLevelNavigationState" : Int, internal
   "StartScreenName" : WString[60], internal
   "DummyTagBool" : Bool, internal
   "DummyTagInt1" : Int, internal
   "DummyTagInt2" : Int, internal
   "DummyTagInt3" : Int, internal
   "DummyDeltaReal" : LReal, internal
   "DummTagReal1" : LReal, internal
   "DummyDeltaInt" : Int, internal
   "MenuInactive" : Int, internal
   "StepNumber" : Int, internal
   "status" : Int AT %DB1.DBW0

text list "Machine State": 0 'Undefined / Kein Job'; 1 'Production / Produktion'; 2 'Startup / Anlauf'; 3 'Paused / Pausiert'; 4 'Stopped / Gestoppt'; 5 'Shutdown / Beenden'; 6 'Undefined / UNBEKANNT'

text list "State": 0 'Off / Aus'; 1 'On / An'

text list "MachineState_Farfield": 0..1 '???'; 1 'OK'; 2 'ERROR / FEHLER'; 3 'PAUSED / HALT'

text list "GroundPos": 0 'No / Nein'; 1 'Yes / Ja'

text list "MachineState": 0 'Kein Job / No Job'; 1 'Produktion / Production'; 2 'Anlauf / Startup'; 3 'Pausiert / Paused'; 4 'Gestoppt / Stopped'; 5 'Beenden / Shutdown'; 6 'Unbekannt / Undefined'

text list "Status": 0 'Man'; 1 'Auto'

text list "Car_color": 3 'Red'; 6 'Blue'; 4 'Green'

text list "MachineStatus": 1 'Busy'; 0 'Idle'; 2 'Run'

text list "MachineMode": 0 'Man'; 1 'Auto'

graphic list "DiagState_3": 0 'DiagOkay_White'; 1 'DiagWarning_White'; 2 'Circle'

graphic list "Machine": 1 'Grafik_Verpackung_Step1_Blink-off'; 2 'Grafik_Verpackung_Step2'; 3 'Grafik_Verpackung_Blink-on'; 6..7 'Grafik_Verpackung_Step1_Blink-off'

graphic list "State": 0..1 'OK'; 3 'Error'

graphic list "CarColorsGraph": 3 'Car_Red'; 6 'Car_Blue_1'; 4 'Car_Green'; 0 'transparent'

